(* Logix 5000 project; controller _GigaDiscovery vendor 1 type 14 code 244 rev 35.11; software revision 35.03; part 21 of 23 *)
(* tags used below, declared in another part *)
   Os : DINT;
   Platform_Open_Cycle_AOI : Sequencer_AOI;
   Timer : TIMER[10];
   All_Rack_Closed_Mem : BOOL;
   DC_Field_Pylon_Motors : UDT_CROUT;   // DC Field Pylon Motors Contactor -Q10101E -Q10103E
   Gondola_Drive_Enable : UDT_CROUT;   // Gondola Drive Ch1-Ch2 Start Enable Contactors -Q16105E -Q16107E
   HMI_Pb_Platform_Open : BOOL;   // HMI Platform Open Command
   HMI_Platform_Close : BOOL;   // HMI Platform Close Command
   I_Compressor_Min_Pressure : BOOL;   // Line Pressure Switch - Minimum Pressure -S21504B
   I_EStop_Pb_OCC1 : UDT_DCI_STOP_TEST;   // +OCC E-stop -S30301F
   I_EStop_Pb_OCC2 : UDT_DCI_STOP_TEST;   // +OCC2 E-Stop -S28502F
   I_Gate_ENTER_G01_Closed : UDT_DCM;   // GATE ENTER (G01) -B25204I
   I_Gate_EXIT_G05_Closed : UDT_DCM;   // GATE EXIT (G05) -B25304I
   I_Gates_Closed : UDT_DCM;   // Gate Closed RFID series -B24802J
   I_OCC1_Stop_Cycle_PB : BOOL;   // Stop Cycle -S30308F
   I_OCC2_ACONFIRM : BOOL;   // OCC2 Allow Main CONFIRM -S28602F
   I_OCC2_Disable : UDT_DCM;   // OCC 2 CONTROL DISABLE Page 310
   I_OCC2_Stop_Cycle_PB : BOOL;   // Stop Cycle -S28606F
   I_OCC_LockOut_Motion : UDT_DCM;   // OCC -Lockout Motion -Q31203E
   I_OCC_Memory_Footpedal : BOOL;
   I_OCC_Operator_Enable_Key : BOOL;   // OCC Console Enabled -S30305F
   I_Operator_Footpedal : BOOL;   // Operator Footpedal -S30901F
   I_Platform_Closed : UDT_DCM;   // Platform Closed RFID Series -B22501J... -B22807J -B22801B
   I_Platform_Line_Min_Pressure_Switch : BOOL;   // Platform Line Minimum Pressure Switch -S21511B
   I_Platform_Opened : UDT_DCM;   // Platform Opened RFID Series -Q23801J -Q23807J
   I_Platform_Pressure_on_Open_Circuit : BOOL;   // Platform Maximum Opening Pressure -S21507B
   I_RESTRAINTS_MainValve_Cosed : BOOL;   // Main Valve Close Limit Switch -B40508I
   I_RESTRAINTS_PressureswitchCompressor : BOOL;   // RESTRAINTS Main Valve Pressure Switch -S40602J
   Mem_All_Rack_Sensor_OFF : BOOL;
   Mem_RESTRAINTS_closed_Correctly : BOOL;
   MODE : BOOL;   // MODE 0 = AUTO 1 = MANUAL -S30801F
   No_Automatic_E_Stop_Cl_0_Request : BOOL;
   No_Automatic_E_Stop_Cl_1_Request : BOOL;
   No_Sfty : Std_to_Sfty;
   O_Close_Platform : BOOL;
   O_Open_Platform : BOOL;
   O_Pilots_Valve_Platform : BOOL;
   O_RESTRAINTS_MainValve : UDT_CROUT;   // Main Valve -B40501I
   Paltform_Cycle_Abborted_Mem : BOOL;   // Paltform Cycle Abborted by Stop Pb Mem
   Pb_Platform_Stop : BOOL;   // Platform Stop Command -S30608F
   Platform_Close_Cycle : Sequencer;
   Platform_CloseMain_Valve_Aux_Comand : BOOL;   // Valvola principale piattaforma QV6515E
   Platform_Open_Cycle : Sequencer;
   Platform_Open_Permissive : Permissive;
   Platform_Open_Permissive_Fail_Edge : DINT;
   Platform_Open_Permissive_Ok : BOOL;
   Platform_OpenMain_Valve_Aux_Comand : BOOL;   // Valvola principale piattaforma QV6515E
   PltaformOpeneded_CycleComplete : BOOL;   // Rilevazione Piattaforme aperte con ciclo Completato
   Power_On_Delay : BOOL;
   ProofTest_Req : BOOL;
   Pylon_Contactor_OFF : BOOL;
   Pylon_Stopped_At_Home : BOOL;   // 5s
   RESTRAINTS_ChA_Open_Memory : BOOL;
   RESTRAINTS_ChB_Open_Memory : BOOL;
   RESTRAINTS_Closed : BOOL;   // All RESTRAINTS Closed
   RESTRAINTS_Rack_Sector_ON : BOOL;
   RESTRAINTS_Sector_Enable_OFF : BOOL;   // ALL RESTRAINTS rack commands OFF
   RESTRAINTS_Unlock_Valve_Pressure : BOOL;
   Start_Platform_AutoCycle_Pylon : BOOL;
   Start_Stop_Cycle : Sequencer;
   Valve_Proof_Test_Cycle : Sequencer;
   Valve_Proof_Test_Ok : BOOL;
(* S_Platform_and_Gates, continued *)

ROUTINE _03_Platform_open_permissive   (* ladder *)
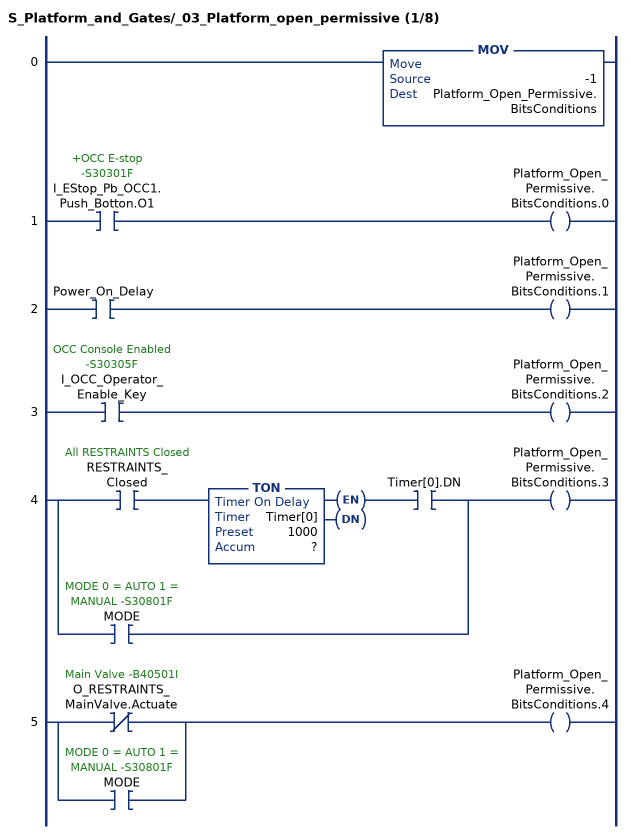
   0: MOV(-1,Platform_Open_Permissive.BitsConditions);
   1: XIC(I_EStop_Pb_OCC1.Push_Botton.O1)OTE(Platform_Open_Permissive.BitsConditions.0);
   2: XIC(Power_On_Delay)OTE(Platform_Open_Permissive.BitsConditions.1);
   3: XIC(I_OCC_Operator_Enable_Key)OTE(Platform_Open_Permissive.BitsConditions.2);
   4: [XIC(RESTRAINTS_Closed) TON(Timer[0],?,?) XIC(Timer[0].DN) ,XIC(MODE) ]OTE(Platform_Open_Permissive.BitsConditions.3);
   5: [XIO(O_RESTRAINTS_MainValve.Actuate) ,XIC(MODE) ]OTE(Platform_Open_Permissive.BitsConditions.4);
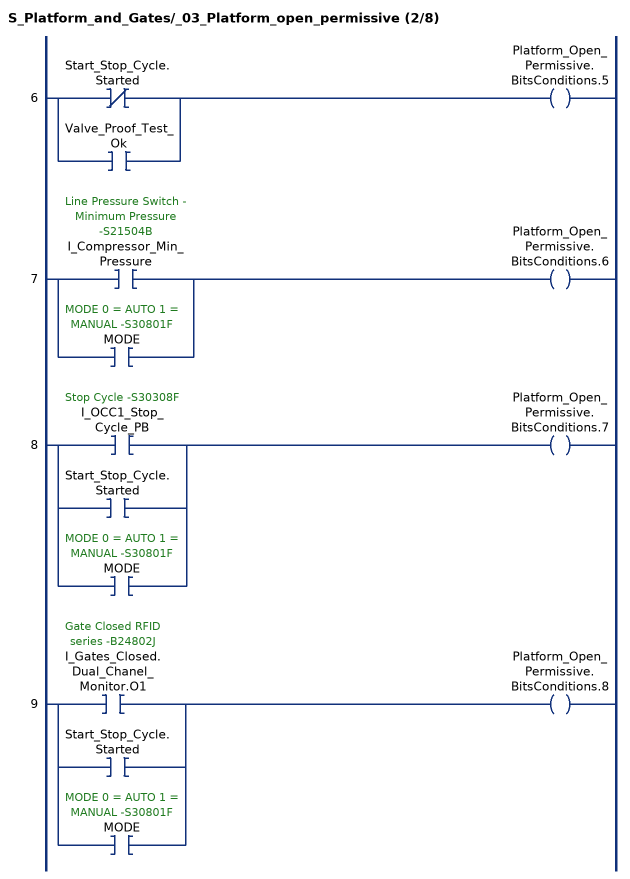
   6: [XIO(Start_Stop_Cycle.Started) ,XIC(Valve_Proof_Test_Ok) ]OTE(Platform_Open_Permissive.BitsConditions.5);
   7: [XIC(I_Compressor_Min_Pressure) ,XIC(MODE) ]OTE(Platform_Open_Permissive.BitsConditions.6);
   8: [XIC(I_OCC1_Stop_Cycle_PB) ,XIC(Start_Stop_Cycle.Started) ,XIC(MODE) ]OTE(Platform_Open_Permissive.BitsConditions.7);
   9: [XIC(I_Gates_Closed.Dual_Chanel_Monitor.O1) ,XIC(Start_Stop_Cycle.Started) ,XIC(MODE) ]OTE(Platform_Open_Permissive.BitsConditions.8);
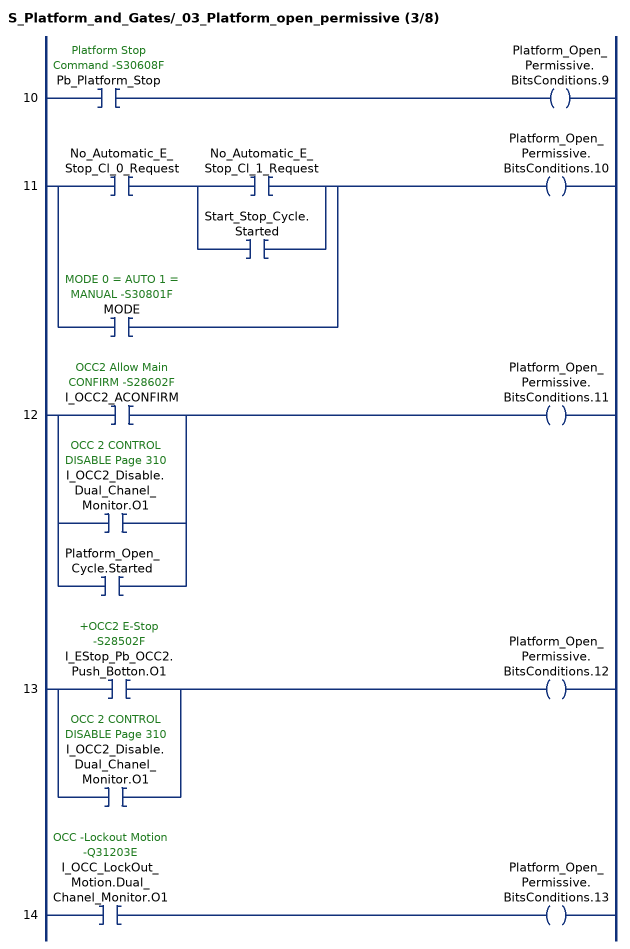
   10: XIC(Pb_Platform_Stop)OTE(Platform_Open_Permissive.BitsConditions.9);
   11: [XIC(No_Automatic_E_Stop_Cl_0_Request) [XIC(No_Automatic_E_Stop_Cl_1_Request) ,XIC(Start_Stop_Cycle.Started) ] ,XIC(MODE) ]OTE(Platform_Open_Permissive.BitsConditions.10);
   12: [XIC(I_OCC2_ACONFIRM) ,XIC(I_OCC2_Disable.Dual_Chanel_Monitor.O1) ,XIC(Platform_Open_Cycle.Started) ]OTE(Platform_Open_Permissive.BitsConditions.11);
   13: [XIC(I_EStop_Pb_OCC2.Push_Botton.O1) ,XIC(I_OCC2_Disable.Dual_Chanel_Monitor.O1) ]OTE(Platform_Open_Permissive.BitsConditions.12);
   14: XIC(I_OCC_LockOut_Motion.Dual_Chanel_Monitor.O1)OTE(Platform_Open_Permissive.BitsConditions.13);
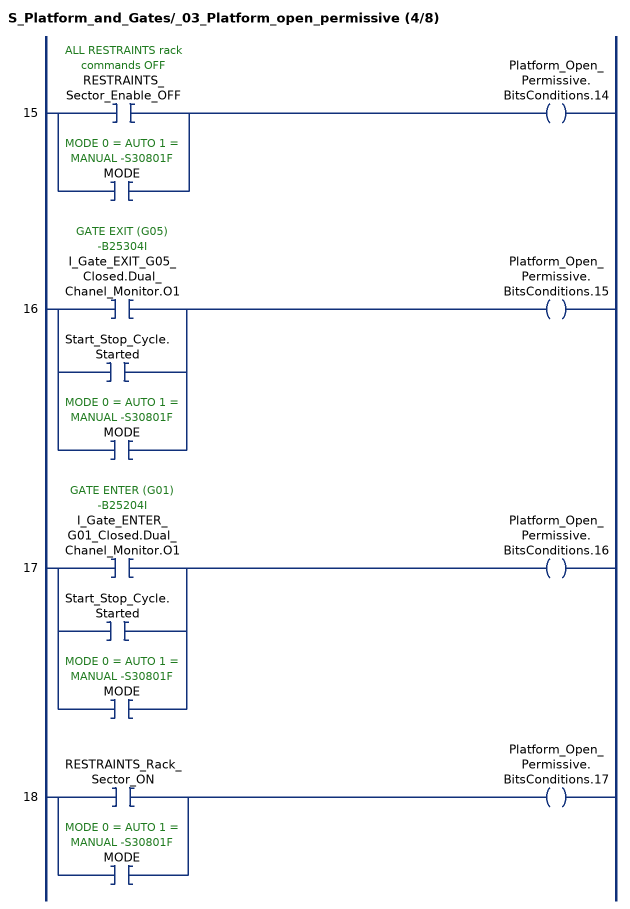
   15: [XIC(RESTRAINTS_Sector_Enable_OFF) ,XIC(MODE) ]OTE(Platform_Open_Permissive.BitsConditions.14);
   16: [XIC(I_Gate_EXIT_G05_Closed.Dual_Chanel_Monitor.O1) ,XIC(Start_Stop_Cycle.Started) ,XIC(MODE) ]OTE(Platform_Open_Permissive.BitsConditions.15);
   17: [XIC(I_Gate_ENTER_G01_Closed.Dual_Chanel_Monitor.O1) ,XIC(Start_Stop_Cycle.Started) ,XIC(MODE) ]OTE(Platform_Open_Permissive.BitsConditions.16);
   18: [XIC(RESTRAINTS_Rack_Sector_ON) ,XIC(MODE) ]OTE(Platform_Open_Permissive.BitsConditions.17);
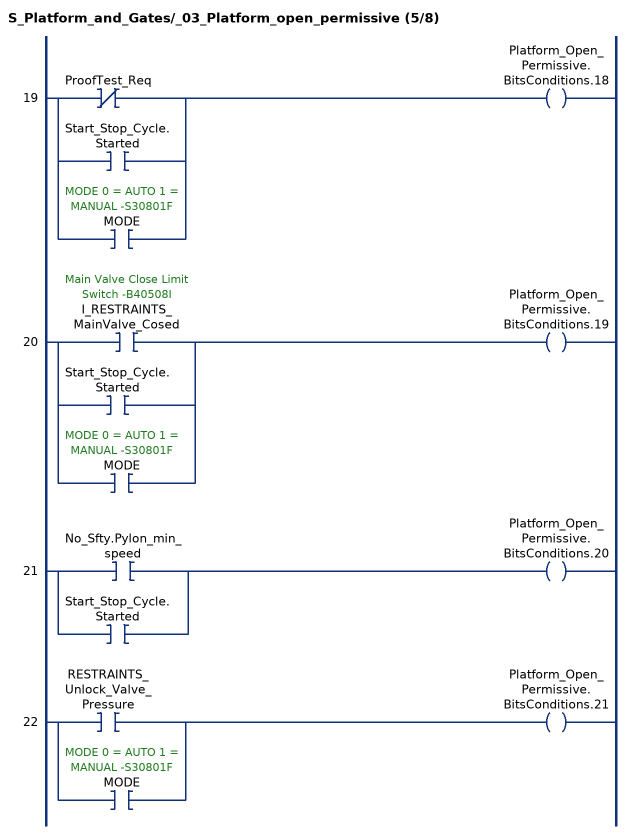
   19: [XIO(ProofTest_Req) ,XIC(Start_Stop_Cycle.Started) ,XIC(MODE) ]OTE(Platform_Open_Permissive.BitsConditions.18);
   20: [XIC(I_RESTRAINTS_MainValve_Cosed) ,XIC(Start_Stop_Cycle.Started) ,XIC(MODE) ]OTE(Platform_Open_Permissive.BitsConditions.19);
   21: [XIC(No_Sfty.Pylon_min_speed) ,XIC(Start_Stop_Cycle.Started) ]OTE(Platform_Open_Permissive.BitsConditions.20);
   22: [XIC(RESTRAINTS_Unlock_Valve_Pressure) ,XIC(MODE) ]OTE(Platform_Open_Permissive.BitsConditions.21);
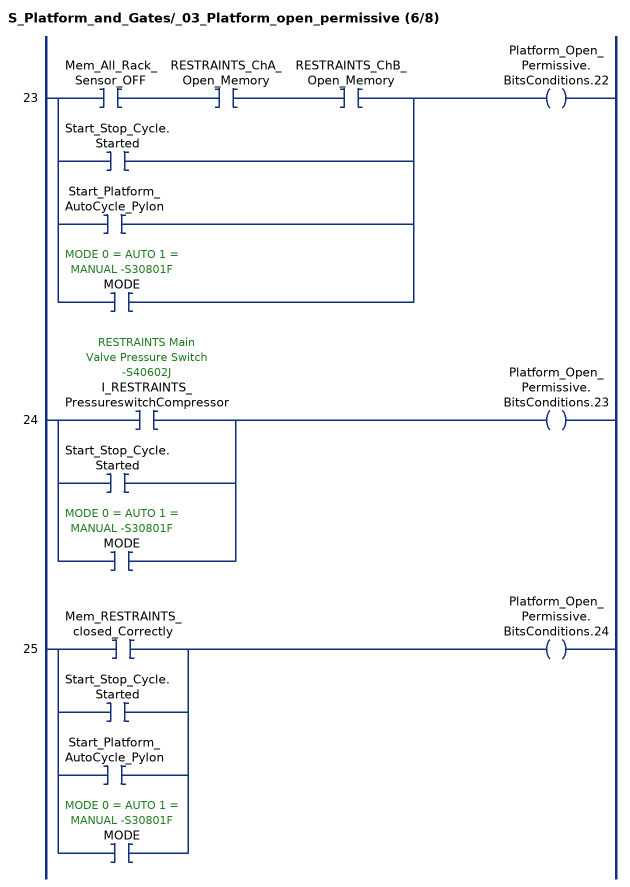
   23: [XIC(Mem_All_Rack_Sensor_OFF) XIC(RESTRAINTS_ChA_Open_Memory) XIC(RESTRAINTS_ChB_Open_Memory) ,XIC(Start_Stop_Cycle.Started) ,XIC(Start_Platform_AutoCycle_Pylon) ,XIC(MODE) ]OTE(Platform_Open_Permissive.BitsConditions.22);
   24: [XIC(I_RESTRAINTS_PressureswitchCompressor) ,XIC(Start_Stop_Cycle.Started) ,XIC(MODE) ]OTE(Platform_Open_Permissive.BitsConditions.23);
   25: [XIC(Mem_RESTRAINTS_closed_Correctly) ,XIC(Start_Stop_Cycle.Started) ,XIC(Start_Platform_AutoCycle_Pylon) ,XIC(MODE) ]OTE(Platform_Open_Permissive.BitsConditions.24);
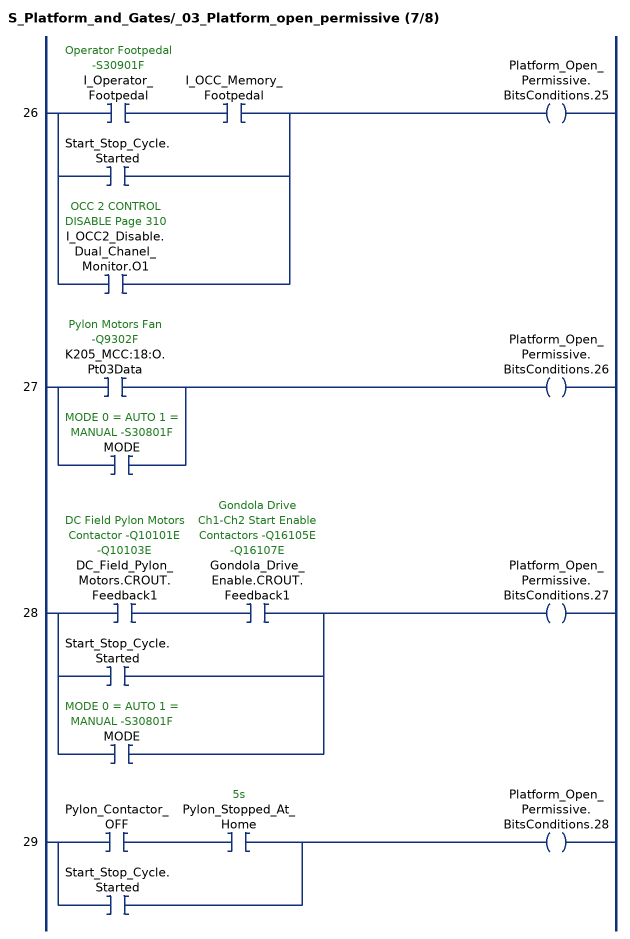
   26: [XIC(I_Operator_Footpedal) XIC(I_OCC_Memory_Footpedal) ,XIC(Start_Stop_Cycle.Started) ,XIC(I_OCC2_Disable.Dual_Chanel_Monitor.O1) ]OTE(Platform_Open_Permissive.BitsConditions.25);
   27: [XIC(K205_MCC:18:O.Pt03Data) ,XIC(MODE) ]OTE(Platform_Open_Permissive.BitsConditions.26);
   28: [XIC(DC_Field_Pylon_Motors.CROUT.Feedback1) XIC(Gondola_Drive_Enable.CROUT.Feedback1) ,XIC(Start_Stop_Cycle.Started) ,XIC(MODE) ]OTE(Platform_Open_Permissive.BitsConditions.27);
   29: [XIC(Pylon_Contactor_OFF) XIC(Pylon_Stopped_At_Home) ,XIC(Start_Stop_Cycle.Started) ]OTE(Platform_Open_Permissive.BitsConditions.28);
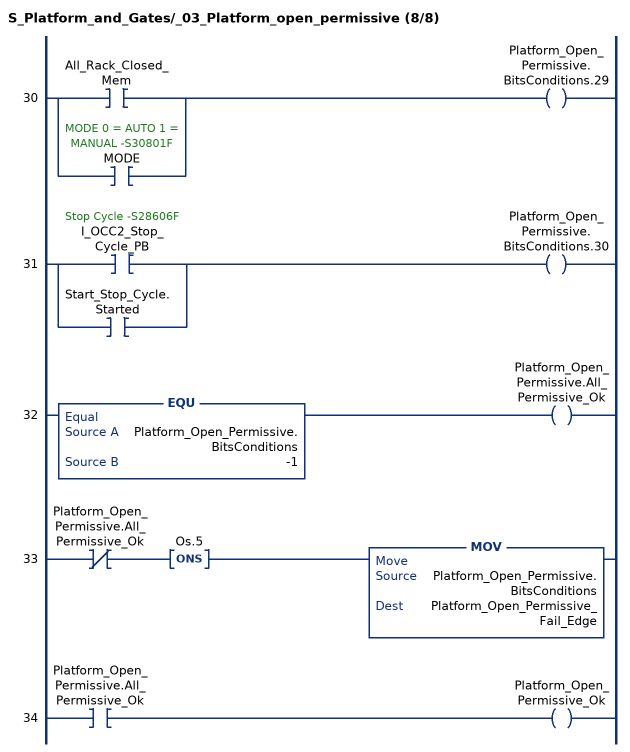
   30: [XIC(All_Rack_Closed_Mem) ,XIC(MODE) ]OTE(Platform_Open_Permissive.BitsConditions.29);
   31: [XIC(I_OCC2_Stop_Cycle_PB) ,XIC(Start_Stop_Cycle.Started) ]OTE(Platform_Open_Permissive.BitsConditions.30);
   32: EQU(Platform_Open_Permissive.BitsConditions,-1)OTE(Platform_Open_Permissive.All_Permissive_Ok);
   33: XIO(Platform_Open_Permissive.All_Permissive_Ok)ONS(Os.5)MOV(Platform_Open_Permissive.BitsConditions,Platform_Open_Permissive_Fail_Edge);
   34: XIC(Platform_Open_Permissive.All_Permissive_Ok)OTE(Platform_Open_Permissive_Ok);
END_ROUTINE

ROUTINE _04_Platform_open_cycle   (* ladder *)
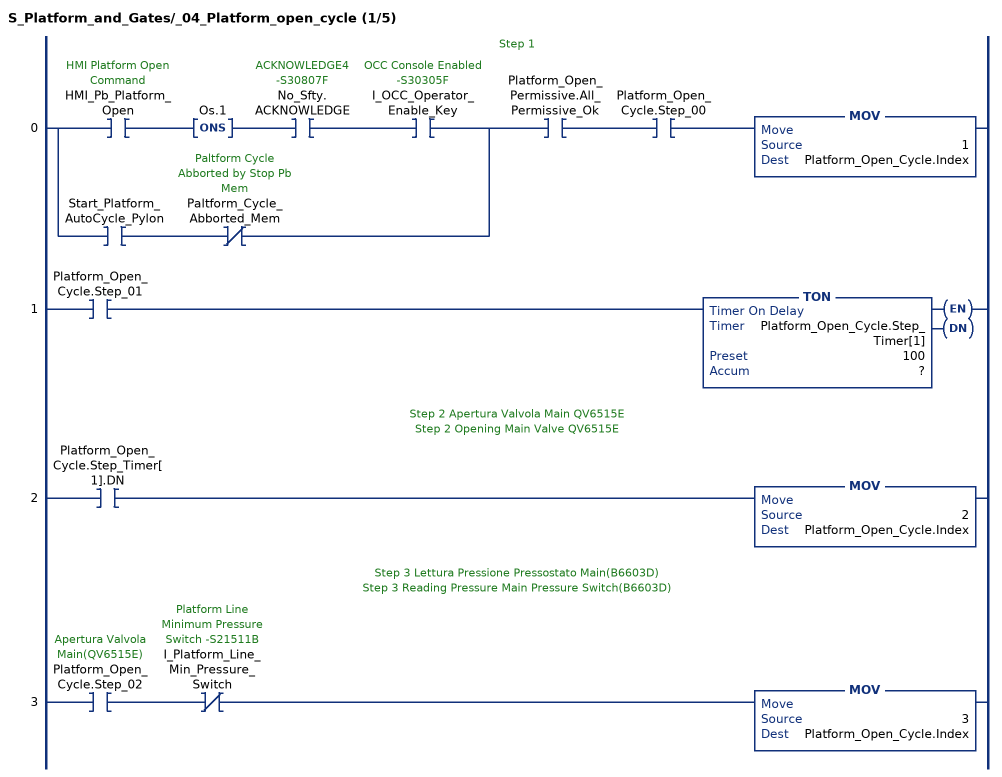
   // Step 1
   0: [XIC(HMI_Pb_Platform_Open) ONS(Os.1) XIC(No_Sfty.ACKNOWLEDGE) XIC(I_OCC_Operator_Enable_Key) ,XIC(Start_Platform_AutoCycle_Pylon) XIO(Paltform_Cycle_Abborted_Mem) ]XIC(Platform_Open_Permissive.All_Permissive_Ok)XIC(Platform_Open_Cycle.Step_00)MOV(1,Platform_Open_Cycle.Index);
   1: XIC(Platform_Open_Cycle.Step_01)TON(Platform_Open_Cycle.Step_Timer[1],?,?);
   // Step 2 Apertura Valvola Main QV6515E
   // Step 2 Opening Main Valve QV6515E
   2: XIC(Platform_Open_Cycle.Step_Timer[1].DN)MOV(2,Platform_Open_Cycle.Index);
   // Step 3 Lettura Pressione Pressostato Main(B6603D)
   // Step 3 Reading Pressure Main Pressure Switch(B6603D)
   3: XIC(Platform_Open_Cycle.Step_02)XIO(I_Platform_Line_Min_Pressure_Switch)MOV(3,Platform_Open_Cycle.Index);
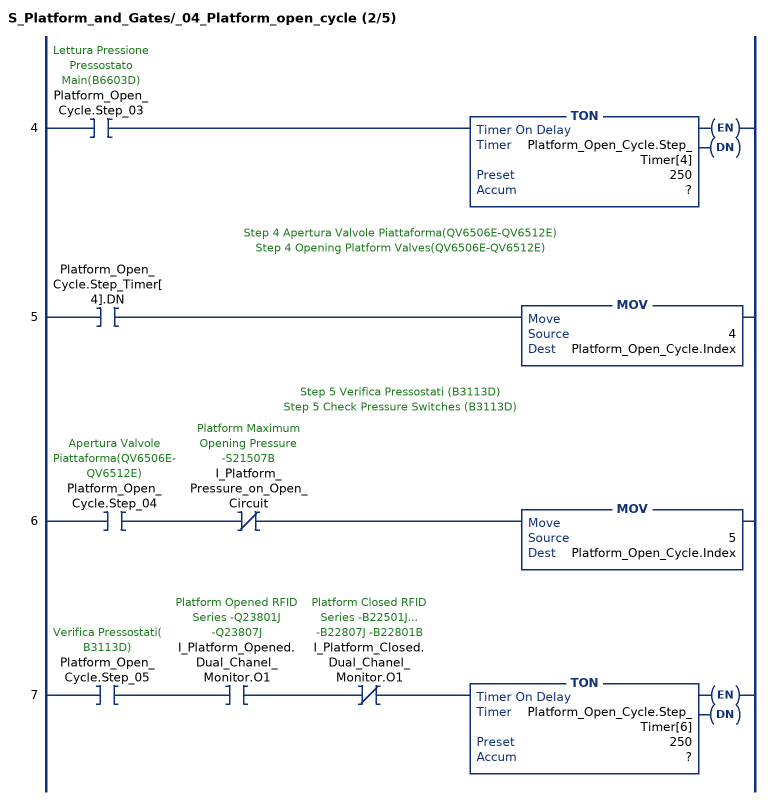
   4: XIC(Platform_Open_Cycle.Step_03)TON(Platform_Open_Cycle.Step_Timer[4],?,?);
   // Step 4 Apertura Valvole Piattaforma(QV6506E-QV6512E)
   // Step 4 Opening Platform Valves(QV6506E-QV6512E)
   5: XIC(Platform_Open_Cycle.Step_Timer[4].DN)MOV(4,Platform_Open_Cycle.Index);
   // Step 5 Verifica Pressostati (B3113D)
   // Step 5 Check Pressure Switches (B3113D)
   6: XIC(Platform_Open_Cycle.Step_04)XIO(I_Platform_Pressure_on_Open_Circuit)MOV(5,Platform_Open_Cycle.Index);
   7: XIC(Platform_Open_Cycle.Step_05)XIC(I_Platform_Opened.Dual_Chanel_Monitor.O1)XIO(I_Platform_Closed.Dual_Chanel_Monitor.O1)TON(Platform_Open_Cycle.Step_Timer[6],?,?);
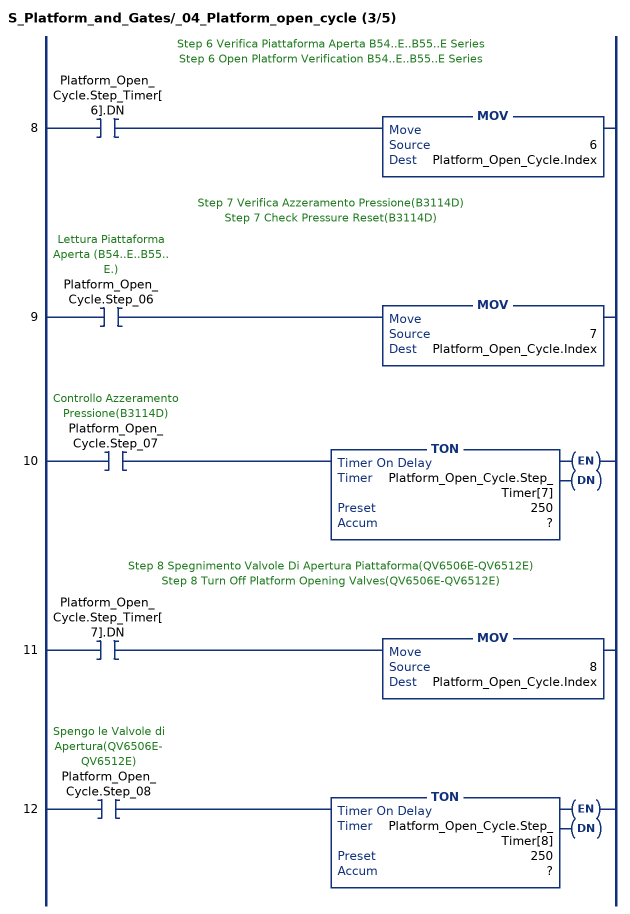
   // Step 6 Verifica Piattaforma Aperta B54..E..B55..E Series
   // Step 6 Open Platform Verification B54..E..B55..E Series
   8: XIC(Platform_Open_Cycle.Step_Timer[6].DN)MOV(6,Platform_Open_Cycle.Index);
   // Step 7 Verifica Azzeramento Pressione(B3114D)
   // Step 7 Check Pressure Reset(B3114D)
   9: XIC(Platform_Open_Cycle.Step_06)MOV(7,Platform_Open_Cycle.Index);
   10: XIC(Platform_Open_Cycle.Step_07)TON(Platform_Open_Cycle.Step_Timer[7],?,?);
   // Step 8 Spegnimento Valvole Di Apertura Piattaforma(QV6506E-QV6512E)
   // Step 8 Turn Off Platform Opening Valves(QV6506E-QV6512E)
   11: XIC(Platform_Open_Cycle.Step_Timer[7].DN)MOV(8,Platform_Open_Cycle.Index);
   12: XIC(Platform_Open_Cycle.Step_08)TON(Platform_Open_Cycle.Step_Timer[8],?,?);
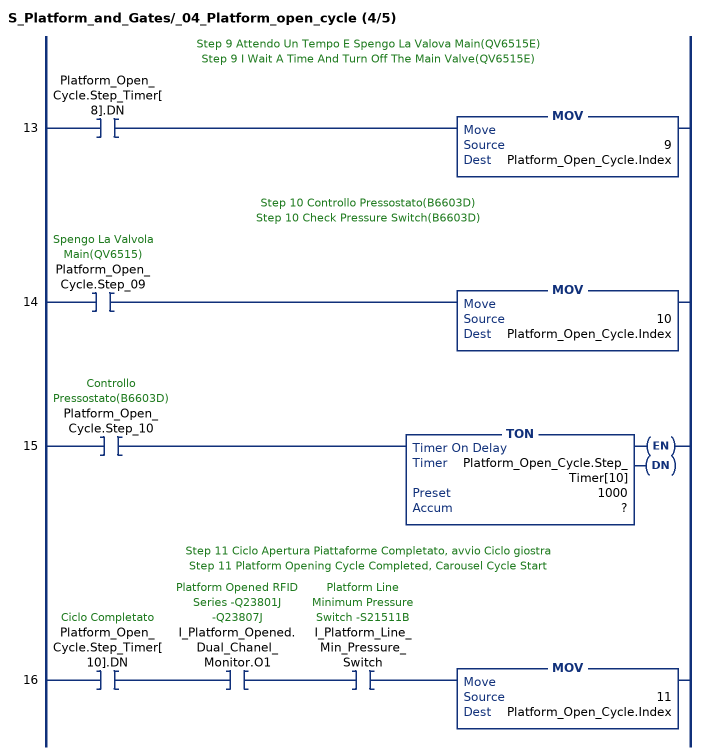
   // Step 9 Attendo Un Tempo E Spengo La Valova Main(QV6515E)
   // Step 9 I Wait A Time And Turn Off The Main Valve(QV6515E)
   13: XIC(Platform_Open_Cycle.Step_Timer[8].DN)MOV(9,Platform_Open_Cycle.Index);
   // Step 10 Controllo Pressostato(B6603D)
   // Step 10 Check Pressure Switch(B6603D)
   14: XIC(Platform_Open_Cycle.Step_09)MOV(10,Platform_Open_Cycle.Index);
   15: XIC(Platform_Open_Cycle.Step_10)TON(Platform_Open_Cycle.Step_Timer[10],?,?);
   // Step 11 Ciclo Apertura Piattaforme Completato, avvio Ciclo giostra
   // Step 11 Platform Opening Cycle Completed, Carousel Cycle Start
   16: XIC(Platform_Open_Cycle.Step_Timer[10].DN)XIC(I_Platform_Opened.Dual_Chanel_Monitor.O1)XIC(I_Platform_Line_Min_Pressure_Switch)MOV(11,Platform_Open_Cycle.Index);
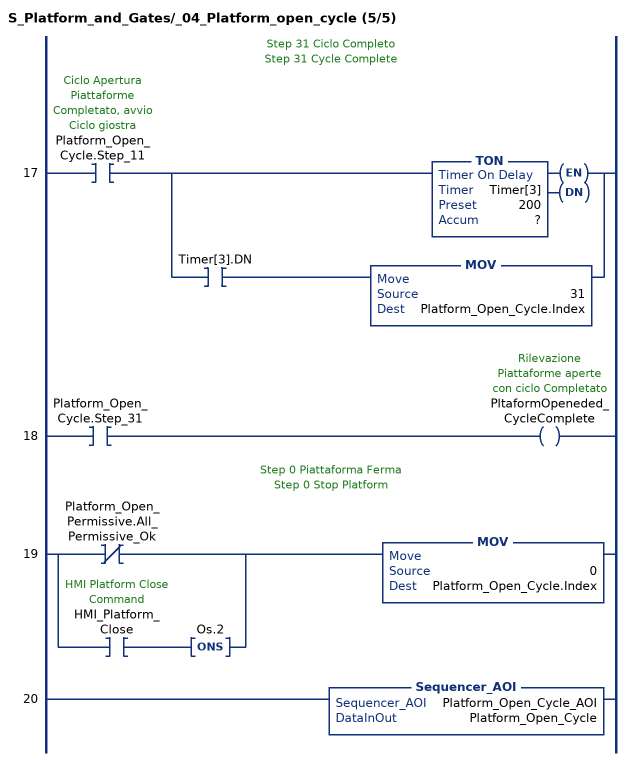
   // Step 31 Ciclo Completo
   // Step 31 Cycle Complete
   17: XIC(Platform_Open_Cycle.Step_11)[TON(Timer[3],?,?) ,XIC(Timer[3].DN) MOV(31,Platform_Open_Cycle.Index) ];
   18: XIC(Platform_Open_Cycle.Step_31)OTE(PltaformOpeneded_CycleComplete);
   // Step 0 Piattaforma Ferma
   // Step 0 Stop Platform
   19: [XIO(Platform_Open_Permissive.All_Permissive_Ok) ,XIC(HMI_Platform_Close) ONS(Os.2) ]MOV(0,Platform_Open_Cycle.Index);
   20: Sequencer_AOI(Platform_Open_Cycle_AOI,Platform_Open_Cycle);
END_ROUTINE

ROUTINE _05_Platform_Stop   (* ladder *)
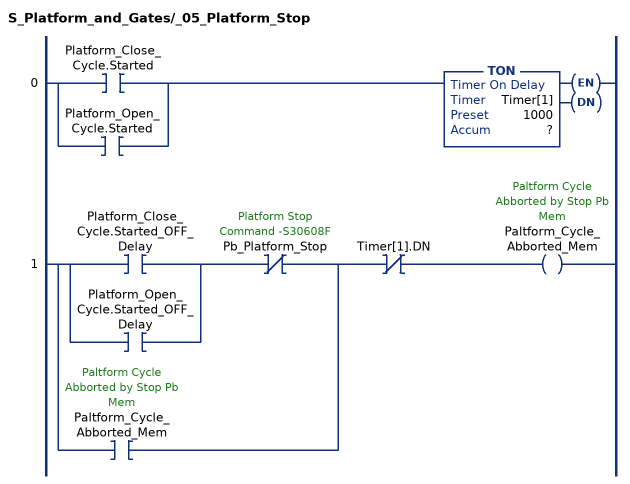
   0: [XIC(Platform_Close_Cycle.Started) ,XIC(Platform_Open_Cycle.Started) ]TON(Timer[1],?,?);
   1: [[XIC(Platform_Close_Cycle.Started_OFF_Delay) ,XIC(Platform_Open_Cycle.Started_OFF_Delay) ] XIO(Pb_Platform_Stop) ,XIC(Paltform_Cycle_Abborted_Mem) ]XIO(Timer[1].DN)OTE(Paltform_Cycle_Abborted_Mem);
END_ROUTINE

ROUTINE _06_Platform_Commands   (* ladder *)
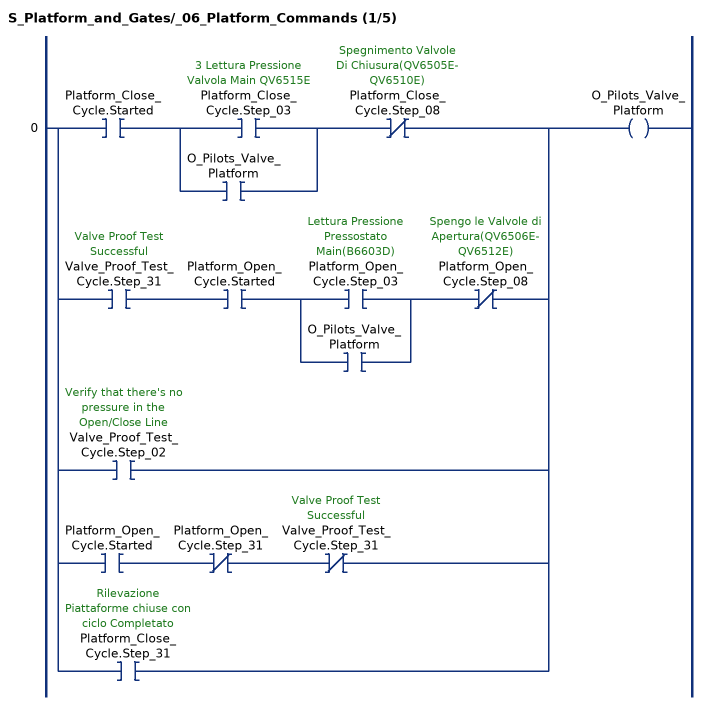
   0: [XIC(Platform_Close_Cycle.Started) [XIC(Platform_Close_Cycle.Step_03) ,XIC(O_Pilots_Valve_Platform) ] XIO(Platform_Close_Cycle.Step_08) ,XIC(Valve_Proof_Test_Cycle.Step_31) XIC(Platform_Open_Cycle.Started) [XIC(Platform_Open_Cycle.Step_03) ,XIC(O_Pilots_Valve_Platform) ] XIO(Platform_Open_Cycle.Step_08) ,XIC(Valve_Proof_Test_Cycle.Step_02) ,XIC(Platform_Open_Cycle.Started) XIO(Platform_Open_Cycle.Step_31) XIO(Valve_Proof_Test_Cycle.Step_31) ,XIC(Platform_Close_Cycle.Step_31) ]OTE(O_Pilots_Valve_Platform);
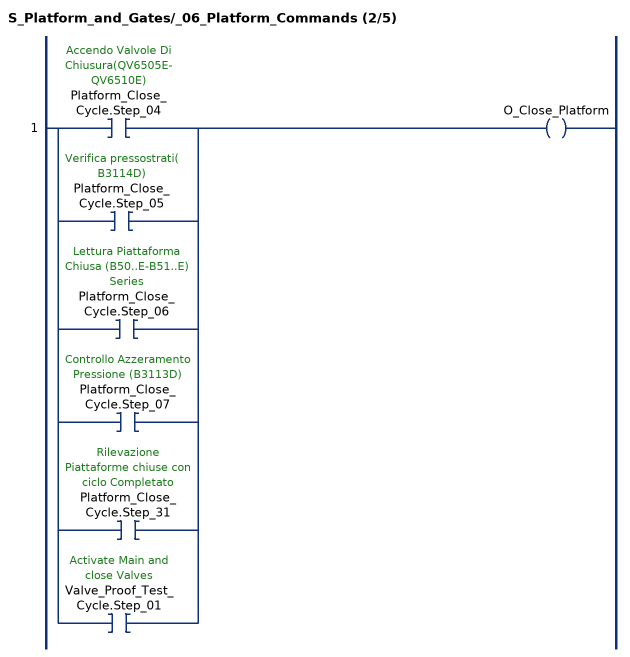
   1: [XIC(Platform_Close_Cycle.Step_04) ,XIC(Platform_Close_Cycle.Step_05) ,XIC(Platform_Close_Cycle.Step_06) ,XIC(Platform_Close_Cycle.Step_07) ,XIC(Platform_Close_Cycle.Step_31) ,XIC(Valve_Proof_Test_Cycle.Step_01) ]OTE(O_Close_Platform);
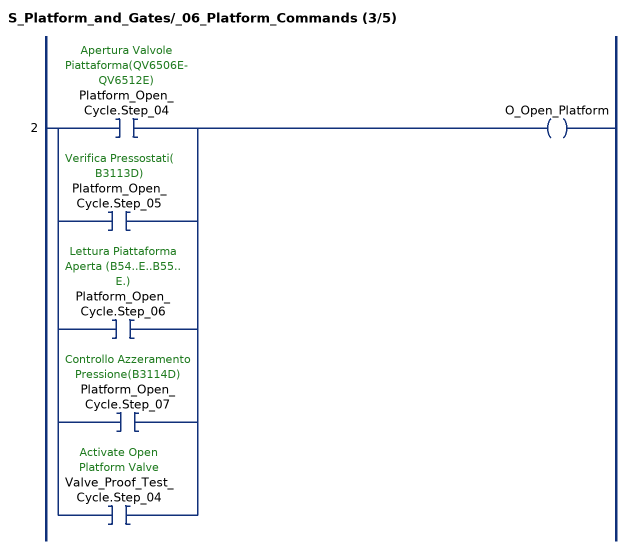
   2: [XIC(Platform_Open_Cycle.Step_04) ,XIC(Platform_Open_Cycle.Step_05) ,XIC(Platform_Open_Cycle.Step_06) ,XIC(Platform_Open_Cycle.Step_07) ,XIC(Valve_Proof_Test_Cycle.Step_04) ]OTE(O_Open_Platform);
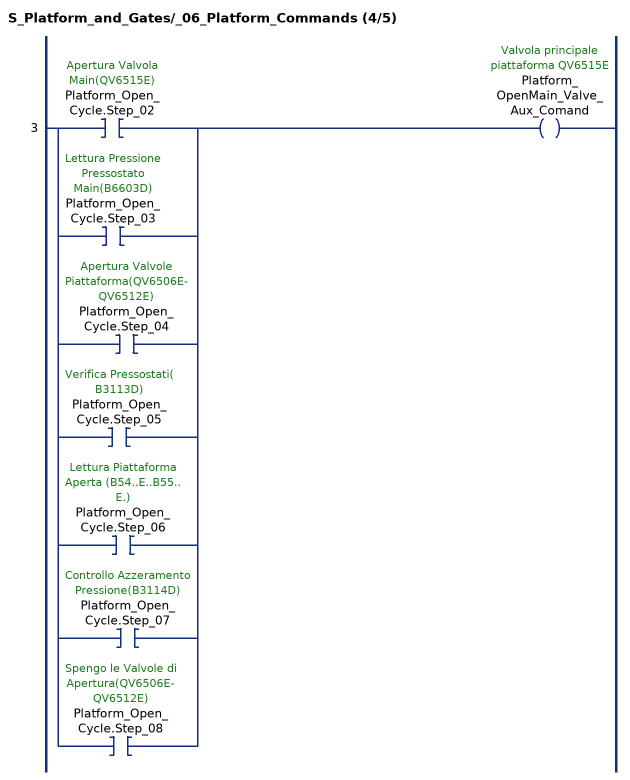
   3: [XIC(Platform_Open_Cycle.Step_02) ,XIC(Platform_Open_Cycle.Step_03) ,XIC(Platform_Open_Cycle.Step_04) ,XIC(Platform_Open_Cycle.Step_05) ,XIC(Platform_Open_Cycle.Step_06) ,XIC(Platform_Open_Cycle.Step_07) ,XIC(Platform_Open_Cycle.Step_08) ]OTE(Platform_OpenMain_Valve_Aux_Comand);
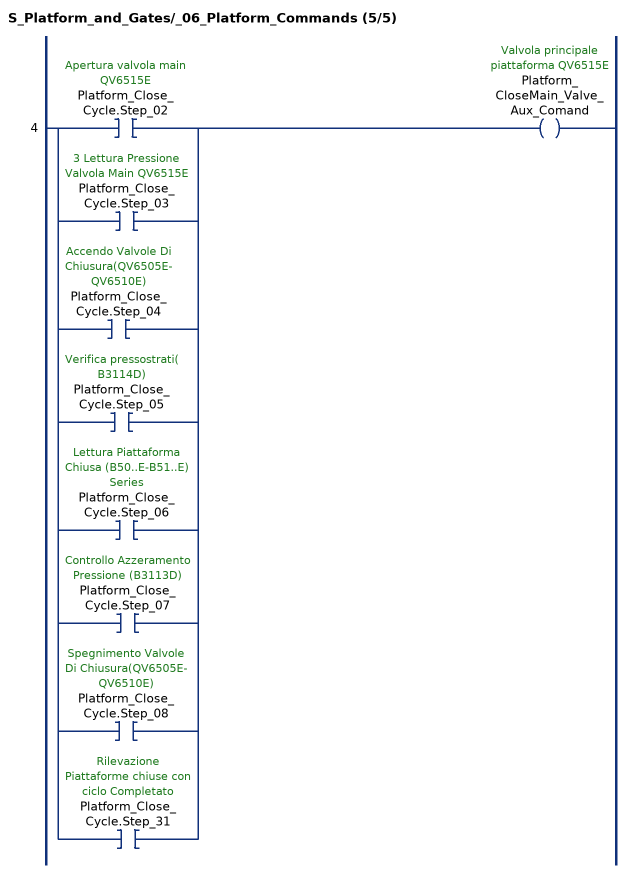
   4: [XIC(Platform_Close_Cycle.Step_02) ,XIC(Platform_Close_Cycle.Step_03) ,XIC(Platform_Close_Cycle.Step_04) ,XIC(Platform_Close_Cycle.Step_05) ,XIC(Platform_Close_Cycle.Step_06) ,XIC(Platform_Close_Cycle.Step_07) ,XIC(Platform_Close_Cycle.Step_08) ,XIC(Platform_Close_Cycle.Step_31) ]OTE(Platform_CloseMain_Valve_Aux_Comand);
END_ROUTINE
